                           END_REGION
                       END_REGION
                       REGION Blad odczytu i awaria zewnetrzna 
                           //zmiana 3.11 word_to_int ze wzgledu na pelny zakres wyjscia przy ujemnym wejsciu
                           "DB331_AI".AI[#i].bSt_Tryb.%X0 := (NOT "DB331_AI".AI[#i].bTrP.%X2) AND (WORD_TO_INT("DB331_AI".AI[#i].wWe) >= 32767 OR WORD_TO_INT("DB331_AI".AI[#i].wWe) <= -32768);
                           "DB331_AI".AI[#i].bSt_Tryb.%X2 := ("DB331_AI".AI[#i].bWeAwrZ AND NOT "DB331_AI".AI[#i].bSt_Tryb.%X12) OR ("DB331_AI".AI[#i].bSym.%X7 AND "DB331_AI".AI[#i].bSt_Tryb.%X12);
                           IF "DB331_AI".AI[#i].bRoZB2.%X0 THEN
                               "DB331_AI".AI[#i].bSt_Tryb.%X0 := 0;
                               "DB331_AI".AI[#i].bSt_Tryb.%X2 := 0;
                           END_IF;
                       END_REGION
                       REGION Przeliczenie wejscia
                           //Z wejscia 
                           IF "DB331_AI".AI[#i].bSt_Tryb.%X14 = 0 THEN
                               "DB331_AI".AI[#i].rWy := (WORD_TO_INT("DB331_AI".AI[#i].wWe) * ("DB331_AI".AI[#i].rZH - "DB331_AI".AI[#i].rZL)) / 27648.0 + "DB331_AI".AI[#i].rZL; //zmiana 3.11 word_to_int
                           ELSE //Zasymulowana, co sekundowa inkrementacja i dekrementacja o zadana wartosc jezeli ustawiony jest ktorys z dwoch bitow
                               IF (("DB331_AI".AI[#i].bSym.%X11 AND "DB331_AI".AI[#i].bSt_Tryb.%X12) OR ("DB331_AI".AI[#i].bWeSymUp AND NOT "DB331_AI".AI[#i].bSt_Tryb.%X12)) AND #Imp_sek THEN
                                   IF "DB331_AI".AI[#i].rWy < "DB331_AI".AI[#i].rZH THEN
                                       "DB331_AI".AI[#i].rWy := "DB331_AI".AI[#i].rWy + "DB331_AI".AI[#i].rSymUp;
                                   ELSE
                                       "DB331_AI".AI[#i].rWy := "DB331_AI".AI[#i].rZH;
                                       ;
                                   END_IF;
                               ELSIF (("DB331_AI".AI[#i].bSym.%X12 AND "DB331_AI".AI[#i].bSt_Tryb.%X12) OR ("DB331_AI".AI[#i].bWeSymDown AND NOT "DB331_AI".AI[#i].bSt_Tryb.%X12)) AND #Imp_sek THEN
                                   IF "DB331_AI".AI[#i].rWy > "DB331_AI".AI[#i].rZL THEN
                                       "DB331_AI".AI[#i].rWy := "DB331_AI".AI[#i].rWy - "DB331_AI".AI[#i].rSymDown;
                                   ELSE
                                       "DB331_AI".AI[#i].rWy := "DB331_AI".AI[#i].rZL;
                                       ;
                                   END_IF;

                                   ;
                               END_IF;
                           END_IF;
                       END_REGION
                       REGION Obsluga awarii zewnetrznej i awarii toru pomiarowego
                           IF "DB331_AI".AI[#i].bSt_Urz = 1 AND "DB331_AI".AI[#i].bAwrUst THEN
                               "DB331_AI".AI[#i].rWy := "DB331_AI".AI[#i].rZL;
                           ELSIF "DB331_AI".AI[#i].bSt_Urz = 1 AND NOT "DB331_AI".AI[#i].bAwrUst THEN
                               "DB331_AI".AI[#i].rWy := "DB331_AI".AI[#i].rZH;
                           END_IF;
                       END_REGION
                       REGION Tryb reczny
                           IF "DB331_AI".AI[#i].bTrP = 4 THEN
                               "DB331_AI".AI[#i].rWy := "DB331_AI".AI[#i].rRoManSter;
                           ELSE
                               "DB331_AI".AI[#i].rRoManSter := "DB331_AI".AI[#i].rWy;
                           END_IF;
                       END_REGION
                       REGION Wyjscie %
                           "DB331_AI".AI[#i].yWy := REAL_TO_INT(100 * ("DB331_AI".AI[#i].rWy - "DB331_AI".AI[#i].rZL) / ("DB331_AI".AI[#i].rZH - "DB331_AI".AI[#i].rZL));
                       END_REGION
                       REGION Sterowanie resetem
                           "DB331_AI".AI[#i].bWyRst := "DB331_AI".AI[#i].bRoZB2.%X0;
                       END_REGION
                       REGION Okreslenie trybu pracy wyjscia
                           IF "DB331_AI".AI[#i].bRoZB1.%X0 THEN
                               "DB331_AI".AI[#i].bTrP := 8;
                           ELSE
                               "DB331_AI".AI[#i].bTrP := 4;
                           END_IF;
                       END_REGION
                       REGION Stan urzadzenia 
                           REGION Przekroczona granica HH pomiaru + filtr
                               IF NOT "DB331_AI".AI[#i].bB.%X0 AND ("DB331_AI".AI[#i].rWy >= "DB331_AI".AI[#i].rGHH) THEN
                                   "DB331_AI".AI[#i].dTmr_HH_Start := true;
                                   ;
                               ELSIF "DB331_AI".AI[#i].rWy < "DB331_AI".AI[#i].rGHH - "DB331_AI".AI[#i].rOffset THEN
                                   "DB331_AI".AI[#i].dTmr_HH_Start := FALSE;
                               END_IF;

                                ;
                               "FC301_Timer"(iTyp := 1,
                                             bOnOff := "DB331_AI".AI[#i].dTmr_HH_Start,
                                             bRst := FALSE,
                                             dCzasZad := "DB331_AI".AI[#i].yCzZadFiltru,
                                             timer_1s := "imp1s",
                                             bOk => "DB331_AI".AI[#i].dTmr_HH_Ok,
                                             dCzasAkt := "DB331_AI".AI[#i].yCzasAktFiltrG);


                           END_REGION
                           REGION Przekroczona granica LL pomiaru + filtr
                               IF NOT "DB331_AI".AI[#i].bB.%X3 AND ("DB331_AI".AI[#i].rWy <= "DB331_AI".AI[#i].rGLL) THEN
                                   "DB331_AI".AI[#i].dTmr_LL_Start := true;
                                   ;
                               ELSIF "DB331_AI".AI[#i].rWy > "DB331_AI".AI[#i].rGLL + "DB331_AI".AI[#i].rFac THEN
                                   "DB331_AI".AI[#i].dTmr_LL_Start := FALSE;
                               END_IF;
                               "FC301_Timer"(iTyp := 1,
                                             bOnOff := "DB331_AI".AI[#i].dTmr_LL_Start,
                                             bRst := FALSE,
                                             dCzasZad := "DB331_AI".AI[#i].yCzZadFiltru,
                                             timer_1s := "imp1s",
                                             bOk => "DB331_AI".AI[#i].dTmr_LL_Ok,
                                             dCzasAkt := "DB331_AI".AI[#i].yCzasAktFiltrD);
                           END_REGION
                           REGION Przypisanie stanow

                               IF "DB331_AI".AI[#i].bSt_Tryb.%X0 OR "DB331_AI".AI[#i].bSt_Tryb.%X2 THEN //Awaria zbiorcza
                                   "DB331_AI".AI[#i].bSt_Urz := 1;
                               ELSIF "DB331_AI".AI[#i].dTmr_HH_Start AND "DB331_AI".AI[#i].dTmr_HH_Ok AND NOT "DB331_AI".AI[#i].bB.%X0 THEN //Awaria HH
                                   "DB331_AI".AI[#i].bSt_Urz := 2;
                               ELSIF "DB331_AI".AI[#i].dTmr_LL_Start AND "DB331_AI".AI[#i].dTmr_LL_Ok AND NOT "DB331_AI".AI[#i].bB.%X3 THEN //Awaria LL
                                   "DB331_AI".AI[#i].bSt_Urz := 32;
                               ELSIF NOT "DB331_AI".AI[#i].bB.%X1 AND ("DB331_AI".AI[#i].rWy >= "DB331_AI".AI[#i].rGH) THEN //Ostrzezenie H
                                   "DB331_AI".AI[#i].bSt_Urz := 4;
                               ELSIF NOT "DB331_AI".AI[#i].bB.%X2 AND ("DB331_AI".AI[#i].rWy <= "DB331_AI".AI[#i].rGL) THEN //Ostrzezenie L
                                   "DB331_AI".AI[#i].bSt_Urz := 16;
                               ELSE //Stan normalnej pracy
                                   "DB331_AI".AI[#i].bSt_Urz := 8;
                               END_IF;

                           END_REGION
                       END_REGION
                       REGION Samokasowanie sygnalow
                           "DB331_AI".AI[#i].bRoZB2 := 0;
                       END_REGION ;

                   END_REGION


              END_IF;
          END_REGION
     END_FOR;
END_FUNCTION

FUNCTION "FC332_AO" : Void   // FC332, SCL
{ S7_Optimized_Access := 'TRUE' }
VERSION : 0.1
   VAR_INPUT
      Nr_Ost_Elementu : Int;   // Numer ostatniego elementu, dla ktorego wykonywana jest klasa
      Nr_Plc : Byte;
   END_VAR
   VAR_TEMP
      i : Int;
   END_VAR
BEGIN
   FOR #i := 1 TO #Nr_Ost_Elementu BY 1 DO
       REGION Opisy bitow sygnalow: bRoz,bSym,bSt,bSt_1,bTrP
           //bRoz - ROZKAZ OPERATORA - DB332.DBW10 - WORD
           //bRozB1
           //"DB332_AO".AO[#i].bRoZB1.%X0 - Tryb pracy: 0-Zdalny reczny; 1-Zdalny auto
           //"DB332_AO".AO[#i].bRoZB1.%X1 - Symulacja wejsc urz: 0-Wylaczona; 1-Zalaczona
           //"DB332_AO".AO[#i].bRoZB1.%X2 - Rezerwa
           //"DB332_AO".AO[#i].bRoZB1.%X3 - Rezerwa
           //"DB332_AO".AO[#i].bRoZB1.%X4 - Rezerwa
           //"DB332_AO".AO[#i].bRoZB1.%X5 - tryb symulacji pomiaru: 1-zalaczony; 2-wylaczony 
           //"DB332_AO".AO[#i].bRoZB1.%X6-X7 - Rezerwa
           //bRozB2 - impulsy  
           //"DB332_AO".AO[#i].bRoZB2.%X0 - Kasuj awarie (impuls)
           //"DB332_AO".AO[#i].bRoZB2.%X1-X7 - Rezerwa (impuls)
           //
           //bSym - SYM WEJSCIA - DB332.DBW12 - WORD
           //"DB332_AO".AO[#i].bSym.%X0 - Aktywacja urz. w systemie (u stawiany tylko z programu)
           //"DB332_AO".AO[#i].bSym.%X1 - Rezerwa
           //"DB332_AO".AO[#i].bSym.%X2-X6 - Rezerwa
           //"DB332_AO".AO[#i].bSym.%X7 - Awaria zewnetrzna: 0-Brak; 1-Aktywny
           //"DB332_AO".AO[#i].bSym.%X8 - Blokada zmiany tr. zdalnego z Auto na Man: 0-Brak; 1-Aktywna
           //"DB332_AO".AO[#i].bSym.%X9-X15 - Rezerwa
           //
           //bSt_Tryb - STAN - DB332.DBW14 - WORD
           //"DB332_AO".AO[#i].bSt_Tryb.%X0 - Awaria toru pomiarowego: 0-Nieaktywna;1-Aktywna
           //"DB332_AO".AO[#i].bSt_Tryb.%X1 - Awaria rezerwa
           //"DB332_AO".AO[#i].bSt_Tryb.%X2 - Awaria zewnetzrna: 0-Nieaktywna; 1-Aktywna
           //"DB332_AO".AO[#i].bSt_Tryb.%X3-X7 - Awaria rezerwa
           //"DB332_AO".AO[#i].bSt_Tryb.%X8 - Urzadzenie aktywowane
           //"DB332_AO".AO[#i].bSt_Tryb.%X9 - Blokada zmaiany tr. zdalnego z Auto na Man: 0-Brak; 1-Aktywna
           //"DB332_AO".AO[#i].bSt_Tryb.%X10-X11 - Awaria rezerwa
           //"DB332_AO".AO[#i].bSt_Tryb.%X12 - Symulacja wejsc urzadzenia: 0-Wylaczona; 1-Zalaczona
           //"DB332_AO".AO[#i].bSt_Tryb.%X13 - Praca z wyjsciami urzadzenia: 0-Wylaczona; 1-Zalaczona
           //"DB332_AO".AO[#i].bSt_Tryb.%X14 - Rezerwa
           //"DB332_AO".AO[#i].bSt_Tryb.%X15 - Stan urzadzenia: 0-Brak odliczania czasu do zamkniecia 1-Odliczanie
           //
           //bSt_Urz - STAN - DB332.DBW16 - INT
           //"DB332_AO".AO[#i].bSt_Urz.%X0 - STAN(1)- Awaria zbiorcza 1-Aktywna; 0-Brak aktywnosci obiektu
           //"DB332_AO".AO[#i].bSt_Urz.%X1 - STAN(2)- Przekroczenie gornej granicy alarmowej
           //"DB332_AO".AO[#i].bSt_Urz.%X2 - STAN(4)- Przekroczenie gornej granicy ostrzegawczej
           //"DB332_AO".AO[#i].bSt_Urz.%X3 - STAN(8)- Urzadzenie: 1-Praca normalne; 0-Inny stan
           //"DB332_AO".AO[#i].bSt_Urz.%X4 - STAN(16)- Prog przekroczenia dolnej granicy ostrzegawczej
           //"DB332_AO".AO[#i].bSt_Urz.%X5 - STAN(32)- Prog przekroczenia dolnej granicy alarmowej
           //"DB332_AO".AO[#i].bSt_Urz.%X6-X7 - STAN- Stan rezerwa
           //
           //bTrP - TRYB PRACY - DB332.DBW17 - INT
           //"DB332_AO".AO[#i].bTrP.%X0 - TRYB PRACY(1): 1-Rezerwa; 0-Brak aktywnosci obiektu
           //"DB332_AO".AO[#i].bTrP.%X1 - Tryb PRACY(2): Rezerwa
           //"DB332_AO".AO[#i].bTrP.%X2 - TRYB PRACY(4) - Tryb Sterowania Zdalnego: 1-Zdalny Reczny; 0-Inny stan
           //"DB332_AO".AO[#i].bTrP.%X3 - TRYB PRACY(8) - Tryb Sterowania Zdalnego: 1-Zdalny Automatyczny; 0-Inny stan
           //"DB332_AO".AO[#i].bTrP.%X4-X7 - Tryb PRACY(16)(32)(64)(128): Rezerwa
           //
           //bL - BLOKADA GENEROWANIA ALARMOW - BYTE
           //"DB332_AO".AO[#i].bB.%X0 - PARAMETR - Blokada generowania alarmu HH: 0-Wylaczona; 1-Zalaczona
           //"DB332_AO".AO[#i].bB.%X1 - PARAMETR - Blokada generowania alarmu H: 0-Wylaczona; 1-Zalaczona
           //"DB332_AO".AO[#i].bB.%X2 - PARAMETR - Blokada generowania alarmu L: 0-Wylaczona; 1-Zalaczona
           //"DB332_AO".AO[#i].bB.%X3 - PARAMETR - Blokada generowania alarmu LL: 0-Wylaczona; 1-Zalaczona
           //"DB332_AO".AO[#i].bB.%X4-X7 - Rezerwa
       END_REGION
      REGION Przepisanie danych do obiektu
          "DB332_AO".AO[#i].yNrID:= #i;
          "DB332_AO".AO[#i].yNrPLC := #Nr_Plc;
                   END_REGION
      REGION Warunek na wykonanie funkcji
          IF "DB332_AO".AO[#i].bWeAkt = 0 THEN //Akcja przy deaktywowaniu obiektu
                  "DB332_AO".AO[#i].bWeAkt := 0;
                  "DB332_AO".AO[#i].bWeAwrZ := 0;
                  "DB332_AO".AO[#i].bWeBlZmAuto := 0;
                  "DB332_AO".AO[#i].bRoZB1 := 0;
                  "DB332_AO".AO[#i].bRoZB2 := 0;
                  "DB332_AO".AO[#i].bSym := 0;
                  "DB332_AO".AO[#i].bSt_Tryb := 0;
                  "DB332_AO".AO[#i].bSt_Urz := 0;
                  "DB332_AO".AO[#i].bTrP := 0;
                  "DB332_AO".AO[#i].bWyRst := 0;

              ELSE
                   REGION Program funkcji
                       REGION Symulacja wejsc - przepisywanie wartosci wejsciowych, gdy nie ma symulacji oprocz bWeAkt
                           IF  "DB332_AO".AO[#i].bSt_Tryb.%X12 = 0 THEN
                               "DB332_AO".AO[#i].bSym.%X7 :=  "DB332_AO".AO[#i].bWeAwrZ;
                               "DB332_AO".AO[#i].bSym.%X8 :=  "DB332_AO".AO[#i].bWeBlZmAuto;
                           END_IF;
                       END_REGION
                       REGION Okreslenie stanow
                           "DB332_AO".AO[#i].bSt_Tryb.%X8 := "DB332_AO".AO[#i].bWeAkt;
                           "DB332_AO".AO[#i].bSt_Tryb.%X9 := (("DB332_AO".AO[#i].bSym.%X8 AND "DB332_AO".AO[#i].bSt_Tryb.%X12) OR ("DB332_AO".AO[#i].bWeBlZmAuto AND NOT "DB332_AO".AO[#i].bSt_Tryb.%X12));
                           "DB332_AO".AO[#i].bSt_Tryb.%X12 := "DB332_AO".AO[#i].bRoZB1.%X1;
                           "DB332_AO".AO[#i].bSt_Tryb.%X14 := "DB332_AO".AO[#i].bRoZB1.%X5;
                           REGION Blokada zmiany trybu zdalny-automatyczny
                               IF "DB332_AO".AO[#i].bSt_Tryb.%X9 AND "DB332_AO".AO[#i].bTrP.%X3 THEN
                                   "DB332_AO".AO[#i].bRoZB1.%X0 := 1;
                               END_IF;
                           END_REGION
                       END_REGION
                       REGION Awaria zewnetrzna
                           IF ("DB332_AO".AO[#i].bWeAwrZ AND NOT "DB332_AO".AO[#i].bSt_Tryb.%X12) OR ("DB332_AO".AO[#i].bSym.%X7 AND "DB332_AO".AO[#i].bSt_Tryb.%X12) THEN
                               "DB332_AO".AO[#i].bSt_Tryb.%X2 := 1;
                           END_IF;
                           IF "DB332_AO".AO[#i].bRoZB2.%X0 THEN
                               "DB332_AO".AO[#i].bSt_Tryb.%X0 := 0;
                               "DB332_AO".AO[#i].bSt_Tryb.%X2 := 0;
                           END_IF;
                       END_REGION
                       REGION Przeliczenie wejscia na rWy i wWy
                           IF "DB332_AO".AO[#i].bTrP=4 THEN 
                               "DB332_AO".AO[#i].rWy := (((("DB332_AO".AO[#i].rZH - "DB332_AO".AO[#i].rZL) / "DB332_AO".AO[#i].rHI_LIM)
                               * "DB332_AO".AO[#i].rFac * "DB332_AO".AO[#i].rRoManSter + "DB332_AO".AO[#i].rZL + "DB332_AO".AO[#i].rOffset) - "DB332_AO".AO[#i].rZL)
                               / ("DB332_AO".AO[#i].rZH - "DB332_AO".AO[#i].rZL)* "DB332_AO".AO[#i].rHI_LIM;
                               "DB332_AO".AO[#i].wWy:=REAL_TO_DINT((("DB332_AO".AO[#i].rZH - "DB332_AO".AO[#i].rZL)/ "DB332_AO".AO[#i].rHI_LIM)*"DB332_AO".AO[#i].rFac*
                                                                   "DB332_AO".AO[#i].rRoManSter+"DB332_AO".AO[#i].rZL+"DB332_AO".AO[#i].rOffset);
                           ELSE
                               "DB332_AO".AO[#i].rWy := (((("DB332_AO".AO[#i].rZH - "DB332_AO".AO[#i].rZL) / "DB332_AO".AO[#i].rHI_LIM)
                               * "DB332_AO".AO[#i].rFac * "DB332_AO".AO[#i].rWe + "DB332_AO".AO[#i].rZL + "DB332_AO".AO[#i].rOffset) - "DB332_AO".AO[#i].rZL)
                               / ("DB332_AO".AO[#i].rZH - "DB332_AO".AO[#i].rZL)* "DB332_AO".AO[#i].rHI_LIM;
                               "DB332_AO".AO[#i].wWy := REAL_TO_DINT((("DB332_AO".AO[#i].rZH - "DB332_AO".AO[#i].rZL) / "DB332_AO".AO[#i].rHI_LIM) * "DB332_AO".AO[#i].rFac *
                                                                     "DB332_AO".AO[#i].rWe + "DB332_AO".AO[#i].rZL + "DB332_AO".AO[#i].rOffset);
                               "DB332_AO".AO[#i].rRoManSter := "DB332_AO".AO[#i].rWy; //Tryb reczny
                           END_IF;
                       END_REGION
                       REGION Obsluga awarii zewnetrznej i awarii toru pomiarowego
                           IF "DB332_AO".AO[#i].bSt_Urz = 1 AND "DB332_AO".AO[#i].bAwrUst THEN
                               "DB332_AO".AO[#i].rWy := "DB332_AO".AO[#i].rZL;
                           ELSIF "DB332_AO".AO[#i].bSt_Urz = 1 AND NOT "DB332_AO".AO[#i].bAwrUst THEN
                               "DB332_AO".AO[#i].rWy := "DB332_AO".AO[#i].rZH;
                           END_IF;
                       END_REGION
                       REGION Wyjscie %
                           "DB332_AO".AO[#i].yWy := REAL_TO_INT("DB332_AO".AO[#i].rWy);
                       END_REGION
                       REGION Sterowanie resetem
                           "DB332_AO".AO[#i].bWyRst :=  "DB332_AO".AO[#i].bRoZB2.%X0;
                       END_REGION
                       REGION Okreslenie trybu pracy wyjscia
                           IF  "DB332_AO".AO[#i].bRoZB1.%X0 THEN
                               "DB332_AO".AO[#i].bTrP := 8;
                           ELSE
                               "DB332_AO".AO[#i].bTrP := 4;
                           END_IF;
                       END_REGION
                       REGION Stan urzadzenia 
                           REGION Przekroczona granica HH pomiaru + filtr
                               "DB332_AO".AO[#i].dTmr_HH_Start := NOT "DB332_AO".AO[#i].bB.%X0 AND ("DB332_AO".AO[#i].rWy >= "DB332_AO".AO[#i].rGHH);
                               "FC301_Timer"(iTyp := 1,
                                             bOnOff := "DB332_AO".AO[#i].dTmr_HH_Start,
                                             bRst := FALSE,
                                             dCzasZad := "DB332_AO".AO[#i].yCzZadFiltru,
                                             timer_1s := "imp1s",
                                             bOk => "DB332_AO".AO[#i].dTmr_HH_Ok,
                                             dCzasAkt := "DB332_AO".AO[#i].yCzasAktFiltrG);


                           END_REGION
                           REGION Przekroczona granica LL pomiaru + filtr
                               "DB332_AO".AO[#i].dTmr_LL_Start := NOT "DB332_AO".AO[#i].bB.%X3 AND ("DB332_AO".AO[#i].rWy <= "DB332_AO".AO[#i].rGLL);
                               "FC301_Timer"(iTyp := 1,
                                             bOnOff := "DB332_AO".AO[#i].dTmr_LL_Start,
                                             bRst := FALSE,
                                             dCzasZad := "DB332_AO".AO[#i].yCzZadFiltru,
                                             timer_1s := "imp1s",
                                             bOk => "DB332_AO".AO[#i].dTmr_LL_Ok,
                                             dCzasAkt := "DB332_AO".AO[#i].yCzasAktFiltrD);
                           END_REGION
                           REGION Przypisanie stanow

                               IF "DB332_AO".AO[#i].bSt_Tryb.%X0 OR "DB332_AO".AO[#i].bSt_Tryb.%X2 THEN //Awaria zbiorcza
                                   "DB332_AO".AO[#i].bSt_Urz := 1;
                               ELSIF "DB332_AO".AO[#i].dTmr_HH_Start AND "DB332_AO".AO[#i].dTmr_HH_Ok AND NOT "DB332_AO".AO[#i].bB.%X0 THEN //Awaria HH
                                   "DB332_AO".AO[#i].bSt_Urz := 2;
                               ELSIF "DB332_AO".AO[#i].dTmr_LL_Start AND "DB332_AO".AO[#i].dTmr_LL_Ok AND NOT "DB332_AO".AO[#i].bB.%X3 THEN //Awaria LL
                                   "DB332_AO".AO[#i].bSt_Urz := 32;
                               ELSIF NOT "DB332_AO".AO[#i].bB.%X1 AND ("DB332_AO".AO[#i].rWy >= "DB332_AO".AO[#i].rGH) THEN //Ostrzezenie H
                                   "DB332_AO".AO[#i].bSt_Urz := 4;
                               ELSIF NOT "DB332_AO".AO[#i].bB.%X2 AND ("DB332_AO".AO[#i].rWy <= "DB332_AO".AO[#i].rGL) THEN //Ostrzezenie L
                                   "DB332_AO".AO[#i].bSt_Urz := 16;
                               ELSE //Stan normalnej pracy
                                   "DB332_AO".AO[#i].bSt_Urz := 8;
                               END_IF;
                           END_REGION
                       END_REGION
                       REGION Samokasowanie sygnalow
                           "DB332_AO".AO[#i].bRoZB2 := 0;
                       END_REGION ;

                   END_REGION


              END_IF;
          END_REGION
     END_FOR;
END_FUNCTION

FUNCTION "FC340_PID" : Void   // FC340, SCL
{ S7_Optimized_Access := 'TRUE' }
VERSION : 0.1
   VAR_INPUT
      Nr_Ost_Elementu : Int;   // Numer ostatniego elementu, dla ktorego wykonywana jest klasa
      Nr_Plc : Byte;
      rCykl : Real;
   END_VAR
   VAR_TEMP
      i : Int;
      Istwert : Real;
      Verstaerk : Real;
      RueckDiff : Real;
      RueckAlt : Real;
      gf : Real;
   END_VAR
   VAR CONSTANT
      Wsp_PV_PER : Real := 0.003616898;   // Wsp uzywany w L137
      Wsp_dLMN : Real := 276.48;   // Wsp uzywany w L302
      Wsp_dLMN_gr : Real := 32511.0;   // Wsp uzywany w L303
      Wsp_dLMN_gr_m : Real := -32512.0;   // Wsp uzywany w L304
   END_VAR
BEGIN
   FOR #i := 1 TO #Nr_Ost_Elementu BY 1 DO
       REGION Opisy bitow sygnalow: bRoz,bSym,bSt,bSt_1,bTrP
           //bRoz - ROZKAZ OPERATORA - DB340.DBW10 - WORD
           //bRozB1
           //"DB340_PID".PID[#i].bRoZB1.%X0 - Trtryb pracy: 0-Zdalny reczny; 1-Zdalny auto
           //"DB340_PID".PID[#i].bRoZB1.%X1 - Symulacja wejsc urz: 0-Wylaczona; 1-Zalaczona
           //"DB340_PID".PID[#i].bRoZB1.%X2 - Rezerwa
           //"DB340_PID".PID[#i].bRoZB1.%X3 - Sterowanie urz. w tr. Zdalnym-Man: 0-Wylacz; 1-Zalacz
           //"DB340_PID".PID[#i].bRoZB1.%X4 - Sterowanie kier. w tr. Zdalnym-Man: 0-Lewa; 1-Prawo
           //"DB340_PID".PID[#i].bRoZB1.%X5 - RoZalSymPom
           //"DB340_PID".PID[#i].bRoZB1.%X6 - Monitoring potwierdzen zal/wyl: 0-Wylaczone; 1-Zalaczone
           //"DB340_PID".PID[#i].bRoZB1.%X7 - Rezerwa
           //bRozB2
           //"DB340_PID".PID[#i].bRoZB2.%X0-X7 - Rezerwa (impuls)
           //
           //bSym - SYM WEJSCIA - DB340.DBW12 - WORD
           //"DB340_PID".PID[#i].bSym.%X0 - Aktywacja urz. w systemie (ustawiany tylko z programu)
           //"DB340_PID".PID[#i].bSym.%X1-X7 - Rezerwa
           //"DB340_PID".PID[#i].bSym.%X8 - Blokada zmiany tr. zdalnego z Auto na Man: 0-Brak; 1-Aktywna
           //"DB340_PID".PID[#i].bSym.%X9-X12 - Rezerwa
           //"DB340_PID".PID[#i].bSym.%X13 - Sledzenie wartosci wejsciowej: 0-Wylaczone; 1-Zalaczone
           //"DB340_PID".PID[#i].bSym.%X14-X15 - Rezerwa
           //
           //bSt_Tryb - STAN - DB340.DBW14 - WORD
           //"DB340_PID".PID[#i].bSt_Tryb.%X0-X7 - Awaria rezerwa
           //"DB340_PID".PID[#i].bSt_Tryb.%X8 - Urzadzenie aktywowane
           //"DB340_PID".PID[#i].bSt_Tryb.%X9 - Blokada zmaiany tr. zdalnego z Auto na Man: 0-Brak; 1-Aktywna
           //"DB340_PID".PID[#i].bSt_Tryb.%X10-X11 - Rezerwa
           //"DB340_PID".PID[#i].bSt_Tryb.%X12 - Symulacja wejsc urzadzenia: 0-Wylaczona; 1-Zalaczona
           //"DB340_PID".PID[#i].bSt_Tryb.%X13 - Rezerwa
           //"DB340_PID".PID[#i].bSt_Tryb.%X14 - StSymPom
           //"DB340_PID".PID[#i].bSt_Tryb.%X15 - Sledzenie sygnalu wejsciowego: 0-Wylaczone; 1-Zalaczone
           //
           //bSt_Urz - STAN - DB340.DBW16 - INT
           //"DB340_PID".PID[#i].bSt_Urz.%X0 - STAN(1)- Rezerwa
           //"DB340_PID".PID[#i].bSt_Urz.%X1 - STAN(2)- Urzadzenie: 1-Wylaczone; 0-Inny stan
           //"DB340_PID".PID[#i].bSt_Urz.%X2 - STAN(4)- Rezerwa
           //"DB340_PID".PID[#i].bSt_Urz.%X3 - STAN(8)- Urzadzenie: 1-Wlaczone; 0-Inny stan
           //"DB340_PID".PID[#i].bSt_Urz.%X4 - STAN(16)- Rezerwa
           //"DB340_PID".PID[#i].bSt_Urz.%X5 - STAN(32)- Rezerwa
           //"DB340_PID".PID[#i].bSt_Urz.%X6-X7 - STAN- Stan rezerwa
           //
           //bTrP - TRYB PRACY - DB340.DBW17 - INT
           //"DB340_PID".PID[#i].bTrP.%X0 - TRYB PRACY(1) - Rezerwa
           //"DB340_PID".PID[#i].bTrP.%X1 - Tryb PRACY(2) - Rezerwa
           //"DB340_PID".PID[#i].bTrP.%X2 - TRYB PRACY(4) - Tryb Sterowania Zdalnego: 1-Zdalny Reczny; 0-Inny stan
           //"DB340_PID".PID[#i].bTrP.%X3 - TRYB PRACY(8) - Tryb Sterowania Zdalnego: 1-Zdalny Automatyczny; 0-Inny stan
           //"DB340_PID".PID[#i].bTrP.%X4-X7 - Tryb PRACY(16)(32)(64)(128): Rezerwa
       END_REGION

       REGION Przepisanie danych do obiektu
           "DB340_PID".PID[#i].yNrID := #i;
           "DB340_PID".PID[#i].yNrPLC := #Nr_Plc;
           "DB340_PID".PID[#i].CYCLE := #rCykl;
       END_REGION

       REGION Warunek na wykonanie funkcji
           IF "DB340_PID".PID[#i].bWeAkt = 0 THEN //Akcja przy deaktywowaniu obiektu
               "DB340_PID".PID[#i].bWeAkt := 0;
               "DB340_PID".PID[#i].bWeZalAuto := 0;
               "DB340_PID".PID[#i].bWeBlZmAuto := 0;
               "DB340_PID".PID[#i].bWeTrck := 0;
               "DB340_PID".PID[#i].bRoZB1 := 0;
               "DB340_PID".PID[#i].bSym := 0;
               "DB340_PID".PID[#i].bSt_Tryb := 0;
               "DB340_PID".PID[#i].bSt_Urz := 0;
               "DB340_PID".PID[#i].bTrP := 0;
               "DB340_PID".PID[#i].bWySter := 0;
               "DB340_PID".PID[#i].QLMN_HLM := 0;
               "DB340_PID".PID[#i].QLMN_LLM := 0;
               "DB340_PID".PID[#i].sbArwHLmOn := 0;
               "DB340_PID".PID[#i].sbArwLLmOn := 0;
               "DB340_PID".PID[#i].LMN := 0;
               "DB340_PID".PID[#i].LMN_PER := 0;
               "DB340_PID".PID[#i].LMN_P := 0;
               "DB340_PID".PID[#i].LMN_I := 0;
               "DB340_PID".PID[#i].LMN_D := 0;
               "DB340_PID".PID[#i].PV := 0;
               "DB340_PID".PID[#i].ER := 0;
               "DB340_PID".PID[#i].sinvAlt := 0;
               "DB340_PID".PID[#i].sIanteilAlt := 0;
               "DB340_PID".PID[#i].sRestInt := 0;
               "DB340_PID".PID[#i].sRestDif := 0; 
               "DB340_PID".PID[#i].sRueck := 0;
               "DB340_PID".PID[#i].sLmn := 0;
           ELSE
               REGION Program funckji
                   REGION Symulacja wejsc - przepisywanie wartosci wejsciowych, gdy nie ma symulacji oprocz bWeAkt
                       IF "DB340_PID".PID[#i].bSt_Tryb.%X12 = 0 THEN
                           "DB340_PID".PID[#i].bSym.%X1 := "DB340_PID".PID[#i].bWeZalAuto;
                           "DB340_PID".PID[#i].bSym.%X8 := "DB340_PID".PID[#i].bWeBlZmAuto;
                           "DB340_PID".PID[#i].bSym.%X13 := "DB340_PID".PID[#i].bWeTrck;
                       END_IF;
                   END_REGION

                   REGION Okreslenie stanow    
                       "DB340_PID".PID[#i].bSt_Tryb.%X8 := "DB340_PID".PID[#i].bWeAkt;
                       "DB340_PID".PID[#i].bSt_Tryb.%X9 := (("DB340_PID".PID[#i].bSym.%X8 AND "DB340_PID".PID[#i].bSt_Tryb.%X12) OR ("DB340_PID".PID[#i].bWeBlZmAuto AND NOT "DB340_PID".PID[#i].bSt_Tryb.%X12));
                       "DB340_PID".PID[#i].bSt_Tryb.%X15 := (("DB340_PID".PID[#i].bSym.%X13 AND "DB340_PID".PID[#i].bSt_Tryb.%X12) OR ("DB340_PID".PID[#i].bWeTrck AND NOT "DB340_PID".PID[#i].bSt_Tryb.%X12));
                       "DB340_PID".PID[#i].bSt_Tryb.%X12 := "DB340_PID".PID[#i].bRoZB1.%X1;
                       "DB340_PID".PID[#i].bSt_Tryb.%X14 := "DB340_PID".PID[#i].bRoZB1.%X5;
                       "DB340_PID".PID[#i].bSt_Urz.%X3 := "DB340_PID".PID[#i].bHlp187;
                       "DB340_PID".PID[#i].bWySter := "DB340_PID".PID[#i].bHlp187;
                       "DB340_PID".PID[#i].bSt_Urz.%X1 :=NOT "DB340_PID".PID[#i].bHlp187;
                   END_REGION
                   REGION Zalaczenie regulatora
                       "DB340_PID".PID[#i].bHlp187 := ("DB340_PID".PID[#i].bTrP.%X3 AND (("DB340_PID".PID[#i].bWeZalAuto AND NOT "DB340_PID".PID[#i].bSt_Tryb.%X12) OR ("DB340_PID".PID[#i].bSym.%X1 AND "DB340_PID".PID[#i].bSt_Tryb.%X12)))
                       OR ("DB340_PID".PID[#i].bTrP.%X2 AND "DB340_PID".PID[#i].bRoZB1.%X3);
                   END_REGION

                   REGION Nadazanie sterowania recznego
                       IF "DB340_PID".PID[#i].bTrP.%X3 THEN
                           "DB340_PID".PID[#i].MAN := "DB340_PID".PID[#i].LMN;
                           "DB340_PID".PID[#i].bRoZB1.%X3 := ("DB340_PID".PID[#i].bWeZalAuto AND NOT "DB340_PID".PID[#i].bSt_Tryb.%X12) OR ("DB340_PID".PID[#i].bSym.%X1 AND "DB340_PID".PID[#i].bSt_Tryb.%X12);
                       END_IF;
                   END_REGION

                   REGION Algorytm PID
                       IF NOT "DB340_PID".PID[#i].bHlp187 THEN
                           "DB340_PID".PID[#i].sIanteilAlt := "DB340_PID".PID[#i].I_ITLVAL;
                           "DB340_PID".PID[#i].LMN := 0;
                           "DB340_PID".PID[#i].QLMN_HLM := 0;
                           "DB340_PID".PID[#i].QLMN_LLM := 0;
                           "DB340_PID".PID[#i].LMN_P := 0;
                           "DB340_PID".PID[#i].LMN_I := 0;
                           "DB340_PID".PID[#i].LMN_D := 0;
                           "DB340_PID".PID[#i].LMN_PER := 0;
                           "DB340_PID".PID[#i].PV := 0;
                           "DB340_PID".PID[#i].ER := 0;
                           "DB340_PID".PID[#i].sinvAlt := 0;
                           "DB340_PID".PID[#i].sRestInt := 0;
                           "DB340_PID".PID[#i].sRestDif := 0;
                           "DB340_PID".PID[#i].sRueck := 0;
                           "DB340_PID".PID[#i].sLmn := 0;
                           "DB340_PID".PID[#i].sbArwHLmOn := 0;
                           "DB340_PID".PID[#i].sbArwLLmOn := 0;

                       ELSE
                           // -----------------------------------------------------------------------------------------------------------------------------------------------
                           #Istwert := INT_TO_REAL(WORD_TO_INT("DB340_PID".PID[#i].PV_PER)) * 100.0 / 27648.0;    // (0-2768 na 0-100)
                           #Istwert := #Istwert * "DB340_PID".PID[#i].PV_FAC + "DB340_PID".PID[#i].PV_OFF;

                           REGION Wybor zrodla PV czy z PV_IN (PVPER=0) czy z PV_PER (PVPER=1)                       
                               IF NOT "DB340_PID".PID[#i].PVPER_ON THEN
                                   #Istwert := "DB340_PID".PID[#i].PV_IN;
                               END_IF;
                           END_REGION

                           "DB340_PID".PID[#i].PV := #Istwert;

                           REGION Wyliczenie uchybu regulacji ErKp=SP_INT-PV
                               "DB340_PID".PID[#i].ErKp := "DB340_PID".PID[#i].SP_INT - "DB340_PID".PID[#i].PV;
                           END_REGION

                           REGION Wyliczenie ER w zaleznosci od ErKp i DEADB_W
                               IF "DB340_PID".PID[#i].ErKp < (- "DB340_PID".PID[#i].DEADB_W) THEN
                                   "DB340_PID".PID[#i].ER := "DB340_PID".PID[#i].ErKp + "DB340_PID".PID[#i].DEADB_W;
                               ELSIF "DB340_PID".PID[#i].ErKp > "DB340_PID".PID[#i].DEADB_W THEN
                                   "DB340_PID".PID[#i].ER := "DB340_PID".PID[#i].ErKp - "DB340_PID".PID[#i].DEADB_W;
                               ELSE
                                   "DB340_PID".PID[#i].ER := 0.0;
                               END_IF;
                           END_REGION

                           REGION Wyznaczenie ErKp
                               "DB340_PID".PID[#i].ErKp := "DB340_PID".PID[#i].ER * "DB340_PID".PID[#i].GAIN;
                           END_REGION

                           REGION Sprawdzenie czy Ti jest mniejsze od polowy cyklu
                               IF "DB340_PID".PID[#i].TI < "DB340_PID".PID[#i].CYCLE * 0.5 THEN
                                   "DB340_PID".PID[#i].TI := "DB340_PID".PID[#i].CYCLE * 0.5;
                               END_IF;
                           END_REGION

                           REGION Sprawdzenie czy Td jest mniejsze od czasu cyklu
                               IF "DB340_PID".PID[#i].TD < "DB340_PID".PID[#i].CYCLE THEN
                                   "DB340_PID".PID[#i].TD := "DB340_PID".PID[#i].CYCLE;
                               END_IF;
                           END_REGION

                           REGION Sprawdzenie czy TmLag jest mniejsze od polowy czasu cyklu 
                               IF "DB340_PID".PID[#i].TM_LAG < "DB340_PID".PID[#i].CYCLE * 0.5 THEN
                                   "DB340_PID".PID[#i].TM_LAG := "DB340_PID".PID[#i].CYCLE * 0.5;
                               END_IF;
                           END_REGION

                           REGION Wyliczenie czesci P 
                               IF "DB340_PID".PID[#i].P_SEL THEN
                                   "DB340_PID".PID[#i].Panteil := "DB340_PID".PID[#i].ErKp;
                               ELSE
                                   "DB340_PID".PID[#i].Panteil := 0.0;
                               END_IF;

                           END_REGION

                           REGION Wyliczanie czesci I
                               IF "DB340_PID".PID[#i].I_SEL
                               THEN
                                   IF "DB340_PID".PID[#i].I_ITL_ON
                                   THEN
                                       "DB340_PID".PID[#i].Ianteil := "DB340_PID".PID[#i].I_ITLVAL;
                                       "DB340_PID".PID[#i].sRestInt := 0.0;
                                   ELSE
                                       IF "DB340_PID".PID[#i].bTrP.%X2 OR "DB340_PID".PID[#i].bSt_Tryb.%X15
                                       THEN
                                           "DB340_PID".PID[#i].Ianteil := "DB340_PID".PID[#i].sLmn - "DB340_PID".PID[#i].Panteil - "DB340_PID".PID[#i].DISV;
                                           "DB340_PID".PID[#i].sRestInt := 0.0;
                                       ELSE
                                           "DB340_PID".PID[#i].Diff := "DB340_PID".PID[#i].CYCLE / "DB340_PID".PID[#i].TI * ("DB340_PID".PID[#i].ErKp + "DB340_PID".PID[#i].sinvAlt) * 0.5 + "DB340_PID".PID[#i].sRestInt;
                                           IF (("DB340_PID".PID[#i].Diff > 0.0) AND "DB340_PID".PID[#i].sbArwHLmOn OR "DB340_PID".PID[#i].INT_HOLD) OR (("DB340_PID".PID[#i].Diff < 0.0) AND "DB340_PID".PID[#i].sbArwLLmOn) THEN
                                               "DB340_PID".PID[#i].Diff := 0.0;
                                           END_IF;
                                           "DB340_PID".PID[#i].Ianteil := "DB340_PID".PID[#i].sIanteilAlt + "DB340_PID".PID[#i].Diff;
                                           "DB340_PID".PID[#i].sRestInt := "DB340_PID".PID[#i].sIanteilAlt - "DB340_PID".PID[#i].Ianteil + "DB340_PID".PID[#i].Diff;
                                       END_IF;
                                   END_IF;
                               ELSE
                                   "DB340_PID".PID[#i].Ianteil := 0.0;
                                   "DB340_PID".PID[#i].sRestInt := 0.0;
                               END_IF;
                           END_REGION

                           REGION Wyliczanie czesci D DO WERYFIKACJI
                               "DB340_PID".PID[#i].Diff := "DB340_PID".PID[#i].ErKp;

                               IF "DB340_PID".PID[#i].bTrP = 4 AND NOT "DB340_PID".PID[#i].D_SEL THEN
                                   #Verstaerk := "DB340_PID".PID[#i].TD / ("DB340_PID".PID[#i].CYCLE * 0.5 + "DB340_PID".PID[#i].TM_LAG);
                                   "DB340_PID".PID[#i].Danteil := ("DB340_PID".PID[#i].Diff - "DB340_PID".PID[#i].sRueck) * #Verstaerk;
                                   #RueckAlt := "DB340_PID".PID[#i].sRueck;
                                   #RueckDiff := "DB340_PID".PID[#i].CYCLE / "DB340_PID".PID[#i].TD * "DB340_PID".PID[#i].Danteil + "DB340_PID".PID[#i].sRestDif;
                                   "DB340_PID".PID[#i].sRueck := #RueckDiff + #RueckAlt;
                                   "DB340_PID".PID[#i].sRestDif := #RueckAlt - "DB340_PID".PID[#i].sRueck + #RueckDiff;
                               ELSE
                                   "DB340_PID".PID[#i].Danteil := 0.0;
                                   "DB340_PID".PID[#i].sRestDif := 0.0;
                                   "DB340_PID".PID[#i].sRueck := "DB340_PID".PID[#i].Diff;
                               END_IF;
                           END_REGION

                           REGION Sumowanie czesci P+I+D i zaklocenia
                               "DB340_PID".PID[#i].dLmn := "DB340_PID".PID[#i].Panteil + "DB340_PID".PID[#i].Ianteil + "DB340_PID".PID[#i].Danteil + "DB340_PID".PID[#i].DISV;
                           END_REGION

                           REGION Tryb sledzenia
                               IF "DB340_PID".PID[#i].bSt_Tryb.%X15 THEN
                                   "DB340_PID".PID[#i].dLmn := "DB340_PID".PID[#i].rTrace;
                                   ;
                               END_IF;
                           END_REGION

                           REGION Tryb pracy zdalnej-recznej i Sprawdzenie ograniczen 
                               IF "DB340_PID".PID[#i].bTrP.%X2 THEN
                                   "DB340_PID".PID[#i].dLmn := "DB340_PID".PID[#i].MAN;
                               ELSE

                                   IF (NOT "DB340_PID".PID[#i].I_ITL_ON) AND "DB340_PID".PID[#i].I_SEL
                                   THEN
                                       IF ("DB340_PID".PID[#i].Ianteil > ("DB340_PID".PID[#i].LMN_HLM - "DB340_PID".PID[#i].DISV)) AND ("DB340_PID".PID[#i].dLmn > "DB340_PID".PID[#i].LMN_HLM) AND (("DB340_PID".PID[#i].dLmn - "DB340_PID".PID[#i].LMN_D) > "DB340_PID".PID[#i].LMN_HLM)
                                       THEN
                                           "DB340_PID".PID[#i].rVal := "DB340_PID".PID[#i].LMN_HLM - "DB340_PID".PID[#i].DISV;
                                           #gf := "DB340_PID".PID[#i].dLmn - "DB340_PID".PID[#i].LMN_HLM;
                                           "DB340_PID".PID[#i].rVal := "DB340_PID".PID[#i].Ianteil - "DB340_PID".PID[#i].rVal;
                                           IF "DB340_PID".PID[#i].rVal > #gf THEN
                                               "DB340_PID".PID[#i].rVal := #gf;
                                           END_IF;
                                           "DB340_PID".PID[#i].Ianteil := "DB340_PID".PID[#i].Ianteil - "DB340_PID".PID[#i].rVal;
                                       ELSE
                                           IF ("DB340_PID".PID[#i].Ianteil < ("DB340_PID".PID[#i].LMN_LLM - "DB340_PID".PID[#i].DISV)) AND ("DB340_PID".PID[#i].dLmn < "DB340_PID".PID[#i].LMN_LLM) AND (("DB340_PID".PID[#i].dLmn - "DB340_PID".PID[#i].LMN_D) < "DB340_PID".PID[#i].LMN_LLM)
                                           THEN
                                               "DB340_PID".PID[#i].rVal := "DB340_PID".PID[#i].LMN_LLM - "DB340_PID".PID[#i].DISV;
                                               #gf := "DB340_PID".PID[#i].dLmn - "DB340_PID".PID[#i].LMN_LLM;
                                               "DB340_PID".PID[#i].rVal := "DB340_PID".PID[#i].Ianteil - "DB340_PID".PID[#i].rVal;
                                               IF "DB340_PID".PID[#i].rVal < #gf THEN
                                                   "DB340_PID".PID[#i].rVal := #gf;
                                               END_IF;
                                               "DB340_PID".PID[#i].Ianteil := "DB340_PID".PID[#i].Ianteil - "DB340_PID".PID[#i].rVal;
                                           END_IF;
                                       END_IF;
                                   END_IF;
                               END_IF;
                           END_REGION

                           "DB340_PID".PID[#i].LMN_P := "DB340_PID".PID[#i].Panteil;
                           "DB340_PID".PID[#i].LMN_I := "DB340_PID".PID[#i].Ianteil;
                           "DB340_PID".PID[#i].LMN_D := "DB340_PID".PID[#i].Danteil;
                           "DB340_PID".PID[#i].sinvAlt := "DB340_PID".PID[#i].ErKp;
                           "DB340_PID".PID[#i].sIanteilAlt := "DB340_PID".PID[#i].Ianteil;
                           "DB340_PID".PID[#i].sbArwHLmOn := 0;
                           "DB340_PID".PID[#i].sbArwLLmOn := 0;
                           IF ("DB340_PID".PID[#i].dLmn >= "DB340_PID".PID[#i].LMN_HLM)
                           THEN
                               "DB340_PID".PID[#i].QLMN_HLM := 1;
                               "DB340_PID".PID[#i].QLMN_LLM := 0;
                               "DB340_PID".PID[#i].dLmn := "DB340_PID".PID[#i].LMN_HLM;
                               "DB340_PID".PID[#i].sbArwHLmOn := 1;
                           ELSE
                               "DB340_PID".PID[#i].QLMN_HLM := 0;
                               IF ("DB340_PID".PID[#i].dLmn <= "DB340_PID".PID[#i].LMN_LLM)
                               THEN
                                   "DB340_PID".PID[#i].QLMN_LLM := 1;
                                   "DB340_PID".PID[#i].dLmn := "DB340_PID".PID[#i].LMN_LLM;
                                   "DB340_PID".PID[#i].sbArwLLmOn := 1;
                               ELSE
                                   "DB340_PID".PID[#i].QLMN_LLM := 0;
                               END_IF;
                           END_IF;
                           "DB340_PID".PID[#i].sLmn := "DB340_PID".PID[#i].dLmn;
                           "DB340_PID".PID[#i].dLmn := "DB340_PID".PID[#i].sLmn * "DB340_PID".PID[#i].LMN_FAC + "DB340_PID".PID[#i].LMN_OFF;
                           "DB340_PID".PID[#i].LMN := "DB340_PID".PID[#i].dLmn;
                           "DB340_PID".PID[#i].dLmn := "DB340_PID".PID[#i].LMN * 2.764800e+002;
                           IF "DB340_PID".PID[#i].dLmn >= 3.251100e+004
                           THEN
                               "DB340_PID".PID[#i].dLmn := 3.251100e+004;
                           ELSE
                               IF "DB340_PID".PID[#i].dLmn <= -3.251200e+004
                               THEN
                                   "DB340_PID".PID[#i].dLmn := -3.251200e+004;
                               END_IF;
                           END_IF;
                           "DB340_PID".PID[#i].LMN_PER := INT_TO_WORD(REAL_TO_INT("DB340_PID".PID[#i].dLmn));

                       END_IF;

                       REGION Okreslenie trybu pracy wyjscia
                           IF NOT "DB340_PID".PID[#i].bRoZB1.%X0 THEN
                               "DB340_PID".PID[#i].bTrP := 4;
                           ELSE
                               "DB340_PID".PID[#i].bTrP := 8;
                           END_IF;
                       END_REGION
                   END_REGION

                   REGION Ustawienia koncowe
                       IF "DB340_PID".PID[#i].bAoff THEN
                           "DB340_PID".PID[#i].bWeZalAuto := 0;
                           ;
                       END_IF;
                   END_REGION
               END_REGION
           END_IF;
       END_REGION
   END_FOR;
END_FUNCTION

FUNCTION "FC352_FF8" : Void   // FC352, SCL
{ S7_Optimized_Access := 'TRUE' }
VERSION : 0.1
   VAR_INPUT
      Nr_Ost_Elementu : Int;   // Numer ostatniego elementu, dla ktorego wykonywana jest klasa
      Nr_Plc : Byte;
      Imp_Sek : Bool;
   END_VAR
   VAR_TEMP
      i : Int;
   END_VAR
BEGIN

   #i := 1;FOR #i := 1 TO #Nr_Ost_Elementu BY 1 DO
      REGION Opisy bitow sygnalow: bRoz,bSym,bSt,bSt_1,bTrP

                       //bRoz - ROZKAZ OPERATORA - DB352.DBW10 - WORD
                       //bRozB1
                       //"DB352_FF8".FF8[#i].bRoZB1.%X0 - Tryb pracy: 0-Zdalny reczny; 1-Zdalny auto
                       //"DB352_FF8".FF8[#i].bRoZB1.%X1 - Symulacja wejsc urz: 0-Wylaczona; 1-Zalaczona
                       //"DB352_FF8".FF8[#i].bRoZB1.%X2 - Rezerwa
                       //"DB352_FF8".FF8[#i].bRoZB1.%X3 - Sterowanie urz. w tr. Zdalnym-Man: 0-Wylacz; 1-Zalacz
                       //"DB352_FF8".FF8[#i].bRoZB1.%X4-X7 - Rezerwa
                       //
                       //bRozB2 - impulsy
                       //"DB332_AO".AO[#i].bRoZB2.%X0-X7 - Rezerwa (impuls)
                       //
                       //bSym - SYM WEJSCIA - DB352.DBW12 - WORD
                       //"DB352_FF8".FF8[#i].bSym.%X0 - Aktywacja urz. w systemie (ustawiany tylko z programu)
                       //"DB352_FF8".FF8[#i].bSym.%X1 - Sterowanie urz. w tr. Zdalnym-Auto: 0-Wylacz; 1-Zalacz
                       //"DB352_FF8".FF8[#i].bSym.%X2-X7 - Rezerwa
                       //"DB352_FF8".FF8[#i].bSym.%X8 - Blokada zmiany tr. zdalnego z Auto na Man: 0-Brak; 1-Aktywna
                       //"DB352_FF8".FF8[#i].bSym.%X9 - Interlock w trybie Zdalnym-Auto: 0-Brak; 1-Aktywny
                       //"DB352_FF8".FF8[#i].bSym.%X10-X15 - Rezerwa
                       //
                       //bSt_Tryb - STAN - DB352.DBW14 - WORD
                       //"DB352_FF8".FF8[#i].bSt_Tryb.%X0-X7
                       //"DB352_FF8".FF8[#i].bSt_Tryb.%X8 - Urzadzenie aktywowane
                       //"DB352_FF8".FF8[#i].bSt_Tryb.%X9 - Blokada zmaiany tr. zdalnego z Auto na Man: 0-Brak; 1-Aktywna
                       //"DB352_FF8".FF8[#i].bSt_Tryb.%X10 - Stan rezerwa
                       //"DB352_FF8".FF8[#i].bSt_Tryb.%X11 - Interlock w trybie Zdalnym-Auto: 0-Brak; 1-Aktywny
                       //"DB352_FF8".FF8[#i].bSt_Tryb.%X12 - Symulacja wejsc urzadzenia: 0-Wylaczona; 1-Zalaczona
                       //"DB352_FF8".FF8[#i].bSt_Tryb.%X13 - Rezerwa
                       //"DB352_FF8".FF8[#i].bSt_Tryb.%X14 - Rezerwa
                       //"DB352_FF8".FF8[#i].bSt_Tryb.%X15 - Rezerwa
                       //
                       //bSt_Urz - STAN - DB352.DBW16 - INT
                       //"DB352_FF8".FF8[#i].bSt_Urz.%X0 - STAN(1)- Awaria zbiorcza 1-Aktywna; 0-Brak aktywnosci obiektu
                       //"DB352_FF8".FF8[#i].bSt_Urz.%X1 - STAN(2)- Urzadzenie: 1-Zamkniete; 0-Inny stan
                       //"DB352_FF8".FF8[#i].bSt_Urz.%X2 - STAN(4)- Rezerwa
                       //"DB352_FF8".FF8[#i].bSt_Urz.%X3 - STAN(8)- Urzadzenie: 1-Otwarte; 0-Inny stan
                       //"DB352_FF8".FF8[#i].bSt_Urz.%X4 - STAN(16)- Rezerwa
                       //"DB352_FF8".FF8[#i].bSt_Urz.%X5 - STAN(32)- Rezerwa
                       //"DB352_FF8".FF8[#i].bSt_Urz.%X6-X7 - STAN(64)(128)- Rezerwa
                       //
                       //bTrP - TRYB PRACY - DB352.DBW17 - INT
                       //"DB352_FF8".FF8[#i].bTrP.%X0 - TRYB PRACY(1) - Rezerwa
                       //"DB352_FF8".FF8[#i].bTrP.%X1 - Tryb PRACY(2) - Rezerwa
                       //"DB352_FF8".FF8[#i].bTrP.%X2 - TRYB PRACY(4) - Tryb Sterowania Zdalnego: 1-Zdalny Reczny; 0-Inny stan
                       //"DB352_FF8".FF8[#i].bTrP.%X3 - TRYB PRACY(8) - Tryb Sterowania Zdalnego: 1-Zdalny Automatyczny; 0-Inny stan
                       //"DB352_FF8".FF8[#i].bTrP.%X4-X7 - Tryb PRACY(16)(32)(64)(128) - Rezerwa
                   END_REGION
      REGION Przepisanie danych do obiektu
          "DB352_FF8".FF8[#i].yNrID := #i;
          "DB352_FF8".FF8[#i].yNrPLC := #Nr_Plc;
                   END_REGION
      REGION Warunek na wykonanie funkcji
          IF "DB352_FF8".FF8[#i].bWeAkt = 0 THEN //Akcja przy deaktywowaniu obiektu
                  "DB352_FF8".FF8[#i].bWeAkt := 0;
                  "DB352_FF8".FF8[#i].bWeZalAuto := 0;
                  "DB352_FF8".FF8[#i].bWeBlZmAuto := 0;
                  "DB352_FF8".FF8[#i].bWeIlock := 0;
                  "DB352_FF8".FF8[#i].bRoZB1 := 0;
                  "DB352_FF8".FF8[#i].bSym := 0;
                  "DB352_FF8".FF8[#i].bSt_Tryb := 0;
                  "DB352_FF8".FF8[#i].bSt_Urz := 0;
                  "DB352_FF8".FF8[#i].bTrP := 0;
                  "DB352_FF8".FF8[#i].bWySter := 0;
                  "DB352_FF8".FF8[#i].dT1_Akt := 0;
                  "DB352_FF8".FF8[#i].dT2_Akt := 0;
                  "DB352_FF8".FF8[#i].dT3_Akt := 0;
                  "DB352_FF8".FF8[#i].iPetle := 0;
                  "DB352_FF8".FF8[#i].bIhlp := 0;
                  "DB352_FF8".FF8[#i].bI1 := 0;
                  "DB352_FF8".FF8[#i].bI2 := 0;
                  "DB352_FF8".FF8[#i].bI3 := 0;
                  "DB352_FF8".FF8[#i].bI4 := 0;
                  "DB352_FF8".FF8[#i].bI5 := 0;
                  "DB352_FF8".FF8[#i].bI6 := 0;
                  "DB352_FF8".FF8[#i].bI7 := 0;
                  "DB352_FF8".FF8[#i].bI8 := 0;
              ELSE